(* Logix 5000 project; controller Seperator 1756-L85E rev 33.11; software revision 33.01; part 3 of 7 *)
(* tags used below, declared in another part *)
   Inp_RunFdbk : BOOL;   // Input Signal: RUN feedback from motor
   Inp_Sim : BOOL;   // 1=Simulate working motor; 0=Start/Stop/ Monitor actual motor
   Inp_OvrdCmd : DINT;   // Override Mode Command: 0=None, 1=Stop, 2=Start
   Cfg_HasRunFdbk : BOOL;   // 1=Motor provides run feedback
   Cfg_UseRunFdbk : BOOL;   // 1=Motor run feedback should be used for failure checking
   Cfg_AllowLocal : BOOL;   // 1=Allow Local Start/Stop without alarm, 0=Start/Stop from HMI/prog only
   Cfg_PCmdClear : ALIAS FOR Mode.Cfg_PCmdClear;
   Cfg_OperStopPrio : BOOL;   // 1=OCmd_Stop available in any mode, 0=OCmd_Stop only in Oper, Maint modes.
   Cfg_ShedOnFailToStart : BOOL;   // 1=Stop Motor and Alarm on Fail to Start; 0=Alarm only on Fail to Start
   PSet_Owner : DINT;   // Program Owner Request ID (non-zero) or Release (zero)
   PCmd_Start : BOOL;   // Program Command to Start Motor
   PCmd_Stop : BOOL;   // Program Command to Stop Motor
   PCmd_Reset : BOOL;   // Program Command to Reset all Alarms requiring Reset
   OCmd_Start : BOOL;   // Operator Command to Start Motor
   OCmd_Stop : BOOL;   // Operator Command to Stop Motor
   OCmd_Bypass : BOOL;   // Operator Command to Bypass all Bypassable Interlocks and Permissives
   OCmd_Check : BOOL;   // Operator Command to Check (not bypass) all Interlocks and Permissives
   MCmd_Disable : BOOL;   // Maintenance Command to Disable Motor
   MCmd_Enable : BOOL;   // Maintenance Command to Enable (allow to run) Motor
   OCmd_Reset : BOOL;   // Operator Command to Reset all Alarms requiring Reset
   OCmd_ResetAckAll : BOOL;   // Operator Command to Reset all Alarms and latched Shed conditions
   Out_Run : BOOL;   // 1=Run Motor, 0=Stop Motor
   Out_Start : BOOL;   // 1=Start Motor, 0=Motor left in current state
   Out_Stop : BOOL;   // 1=Stop Motor, 0=Motor left in current state
   Val_Cmd : SINT;   // Device Command 0=None, 1=Stop, 2=Start
   Val_Fdbk : SINT;   // Device Feedback 0=Stopped, 1=Running
   Val_Sts : SINT;   // Device Confirmed Sts 0=? 1=Stopped, 2=Running, 7=Stopping, 8=Starting, 33=Disabled
   Val_Fault : SINT;   // Device Fault Status 0=None, 16=Fail to Start, 17 = Fail to Stop, 32=I/O Fault, 34=Config Error
   Val_Owner : DINT;   // Current Object Owner ID (0=not owned)
   Val_Notify : SINT;   // Current Alarm Level and Acknowledgement (enumeration)
   Sts_Stopped : BOOL;   // 1=Motor requested to stop and is confirmed stopped
   Sts_Starting : BOOL;   // 1=Motor requested to run and awaiting run feedback
   Sts_Running : BOOL;   // 1=Motor requested to run and is confirmed running
   Sts_Stopping : BOOL;   // 1=Motor requested to stop and awaiting stopped feedback
   Sts_Available : BOOL;   // 1=Motor available for control by automation (Prog)
   Sts_Disabled : BOOL;   // 1=Motor is Disabled
   Sts_NotRdy : BOOL;   // 1=Motor is Not Ready to Run (independent of Mode)
   Sts_AlmInh : BOOL;   // 1=An Alarm is Shelved, Disabled or Suppressed: display icon
   Sts_Err : BOOL;   // 1=Error in Config: see detail bits for reason
   Sts_Hand : ALIAS FOR Mode.Sts_Hand;
   Sts_Maint : ALIAS FOR Mode.Sts_Maint;
   Sts_Ovrd : ALIAS FOR Mode.Sts_Ovrd;
   Sts_Prog : ALIAS FOR Mode.Sts_Prog;
   Sts_Oper : ALIAS FOR Mode.Sts_Oper;
   Sts_FailToStart : ALIAS FOR FailToStart.Inp;   // 1=Motor Failed to Start (one-shot)
   Sts_FailToStop : ALIAS FOR FailToStop.Inp;   // 1=Motor Failed to Stop
   Sts_IOFault : ALIAS FOR IOFault.Inp;   // I/O Comm Fault Status (0=OK, 1=Bad)
   Rdy_Start : BOOL;   // 1=Ready to receive OCmd_Start (enables HMI button)
   Rdy_Stop : BOOL;   // 1=Ready to receive OCmd_Stop (enables HMI button)
   Rdy_Reset : BOOL;   // 1=At least one Alarm or Latched Shed requires Reset
   Rdy_ResetAckAll : BOOL;   // 1=At least one Alarm or latched Shed condition requires Reset or Ack
   P_Motor : BOOL;   // Unique Parameter Name for auto - discovery
   Mode : P_Mode;   // Motor Mode Selection
   IOFault : P_Alarm;   // I/O Fault Alarm
   IntlkTrip : P_Alarm;   // Interlock Trip Alarm
   FailToStop : P_Alarm;   // Motor Failed to Stop Alarm
   FailToStart : P_Alarm;   // Motor Failed to Start Alarm
   Wrk_Run : BOOL;   // 1=Motor should be "running", 0=should be "stopped"
   Wrk_SimRunT : TIMER;   // Simulation Delay until Running
   Wrk_StopT : TIMER;   // Stop Check Timer
   Wrk_StartT : TIMER;   // Start Check Timer
   Wrk_SimStopT : TIMER;   // Simulation Delay until Stopped
   Wrk_RunFdbk : BOOL;   // Run Feedback based on mode, simulation, etc. 1=running
   Wrk_Notify : DINT;   // Buffer for building Val_Notify
   Wrk_Cmd : SINT;   // Buffer for building Val_Cmd
   Wrk_Sts : SINT;   // Buffer for building Val_Sts
   Wrk_Fault : SINT;   // Buffer for building Val_Fault
   Wrk_Retrigger : BOOL;   // Maint Start issued while running or Stop while stopped
   Wrk_FailToStart : BOOL;   // Fail to Start Fault (latched) stops motor and requires reset
   Wrk_IOFault : BOOL;   // I/O Fault (latched) stops motor and requires reset
   Starting : SFC_STEP;
   Stopped : SFC_STEP;
   Stopping : SFC_STEP;
(* P_Motor, continued *)

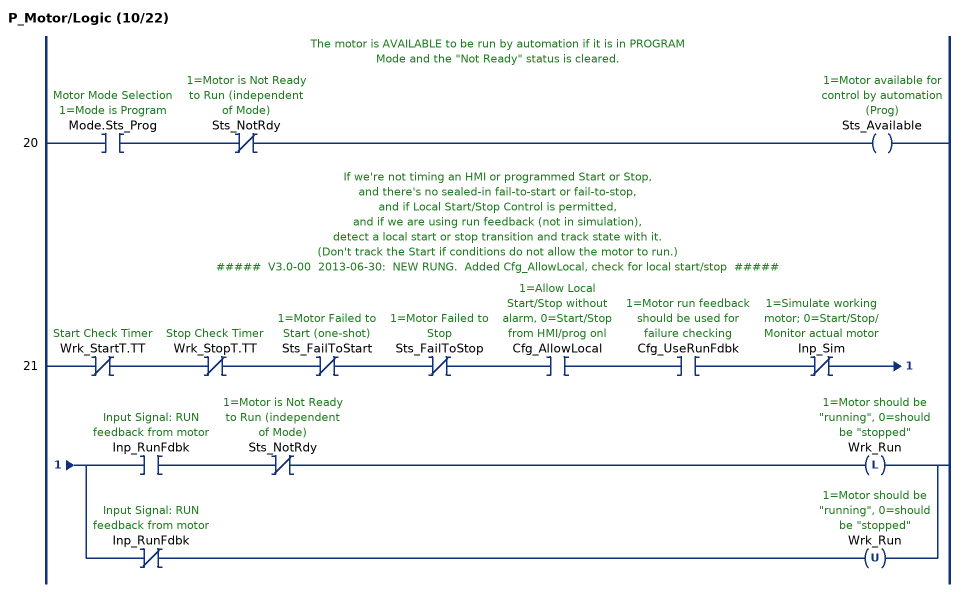
   // The motor is AVAILABLE to be run by automation if it is in PROGRAM
   // Mode and the "Not Ready" status is cleared.
   20: XIC(Mode.Sts_Prog)XIO(Sts_NotRdy)OTE(Sts_Available);
   // If we're not timing an HMI or programmed Start or Stop,
   // and there's no sealed-in fail-to-start or fail-to-stop,
   // and if Local Start/Stop Control is permitted,
   // and if we are using run feedback (not in simulation),
   // detect a local start or stop transition and track state with it.
   // (Don't track the Start if conditions do not allow the motor to run.)
   // #####  V3.0-00  2013-06-30:  NEW RUNG.  Added Cfg_AllowLocal, check for local start/stop  #####
   21: XIO(Wrk_StartT.TT)XIO(Wrk_StopT.TT)XIO(Sts_FailToStart)XIO(Sts_FailToStop)XIC(Cfg_AllowLocal)XIC(Cfg_UseRunFdbk)XIO(Inp_Sim)[XIC(Inp_RunFdbk) XIO(Sts_NotRdy) OTL(Wrk_Run) ,XIO(Inp_RunFdbk) OTU(Wrk_Run) ];
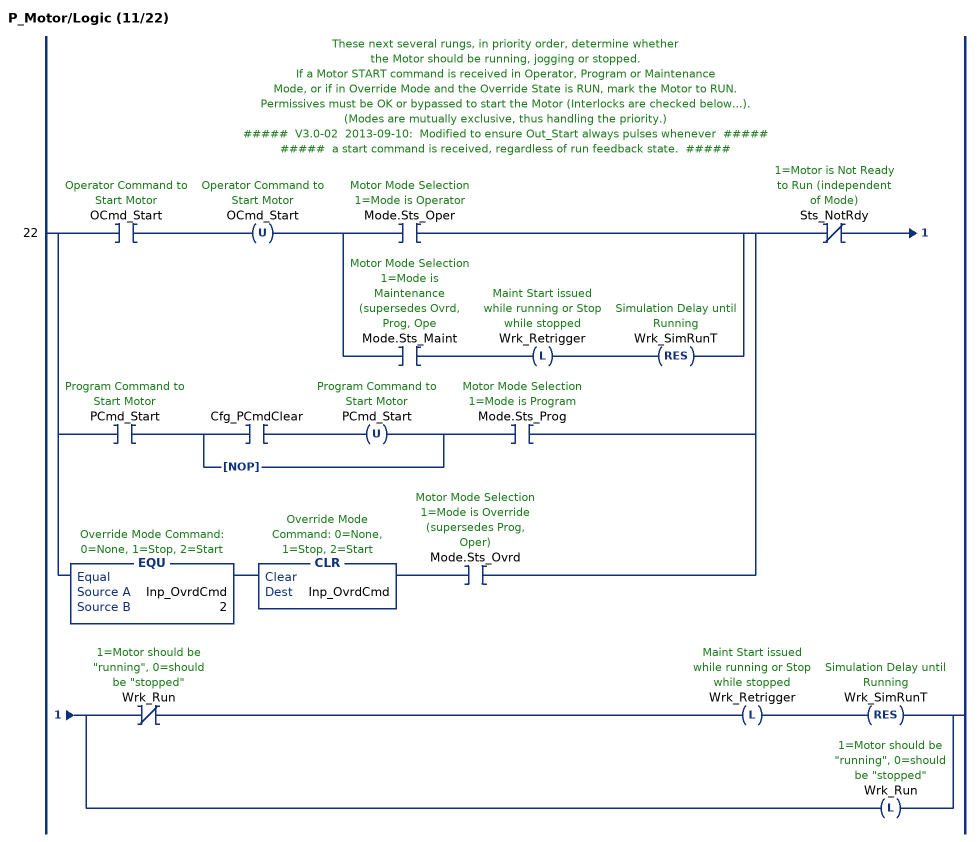
   // These next several rungs, in priority order, determine whether
   // the Motor should be running, jogging or stopped.
   // If a Motor START command is received in Operator, Program or Maintenance
   // Mode, or if in Override Mode and the Override State is RUN, mark the Motor to RUN.
   // Permissives must be OK or bypassed to start the Motor (Interlocks are checked below...).
   // (Modes are mutually exclusive, thus handling the priority.)
   // #####  V3.0-02  2013-09-10:  Modified to ensure Out_Start always pulses whenever  #####
   // #####  a start command is received, regardless of run feedback state.  #####
   22: [XIC(OCmd_Start) OTU(OCmd_Start) [XIC(Mode.Sts_Oper) ,XIC(Mode.Sts_Maint) OTL(Wrk_Retrigger) RES(Wrk_SimRunT) ] ,XIC(PCmd_Start) [XIC(Cfg_PCmdClear) OTU(PCmd_Start) ,NOP() ] XIC(Mode.Sts_Prog) ,EQU(Inp_OvrdCmd,2) CLR(Inp_OvrdCmd) XIC(Mode.Sts_Ovrd) ]XIO(Sts_NotRdy)[XIO(Wrk_Run) OTL(Wrk_Retrigger) RES(Wrk_SimRunT) ,OTL(Wrk_Run) ];
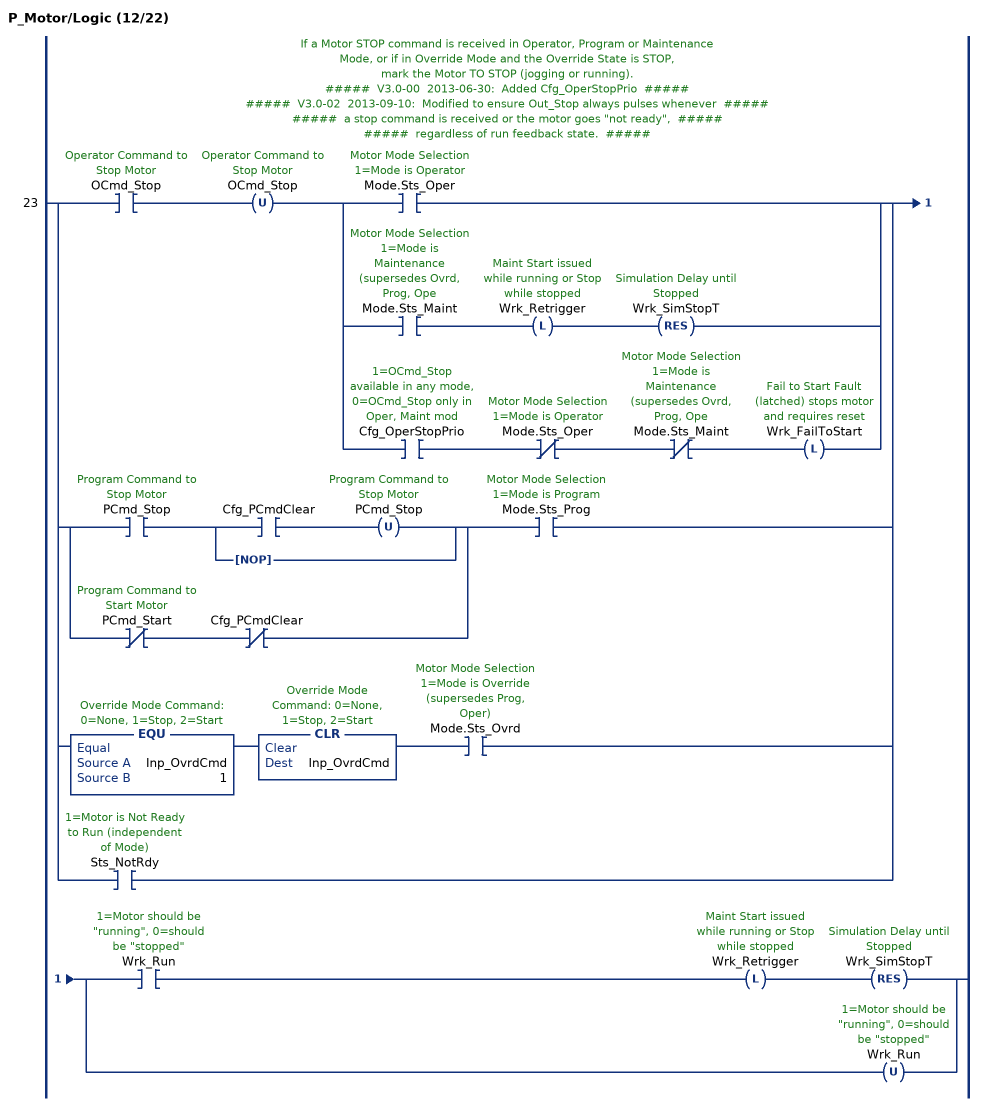
   // If a Motor STOP command is received in Operator, Program or Maintenance
   // Mode, or if in Override Mode and the Override State is STOP,
   // mark the Motor TO STOP (jogging or running).
   // #####  V3.0-00  2013-06-30:  Added Cfg_OperStopPrio  #####
   // #####  V3.0-02  2013-09-10:  Modified to ensure Out_Stop always pulses whenever  #####
   // #####  a stop command is received or the motor goes "not ready",  #####
   // #####  regardless of run feedback state.  #####
   23: [XIC(OCmd_Stop) OTU(OCmd_Stop) [XIC(Mode.Sts_Oper) ,XIC(Mode.Sts_Maint) OTL(Wrk_Retrigger) RES(Wrk_SimStopT) ,XIC(Cfg_OperStopPrio) XIO(Mode.Sts_Oper) XIO(Mode.Sts_Maint) OTL(Wrk_FailToStart) ] ,[XIC(PCmd_Stop) [XIC(Cfg_PCmdClear) OTU(PCmd_Stop) ,NOP() ] ,XIO(PCmd_Start) XIO(Cfg_PCmdClear) ] XIC(Mode.Sts_Prog) ,EQU(Inp_OvrdCmd,1) CLR(Inp_OvrdCmd) XIC(Mode.Sts_Ovrd) ,XIC(Sts_NotRdy) ][XIC(Wrk_Run) OTL(Wrk_Retrigger) RES(Wrk_SimStopT) ,OTU(Wrk_Run) ];
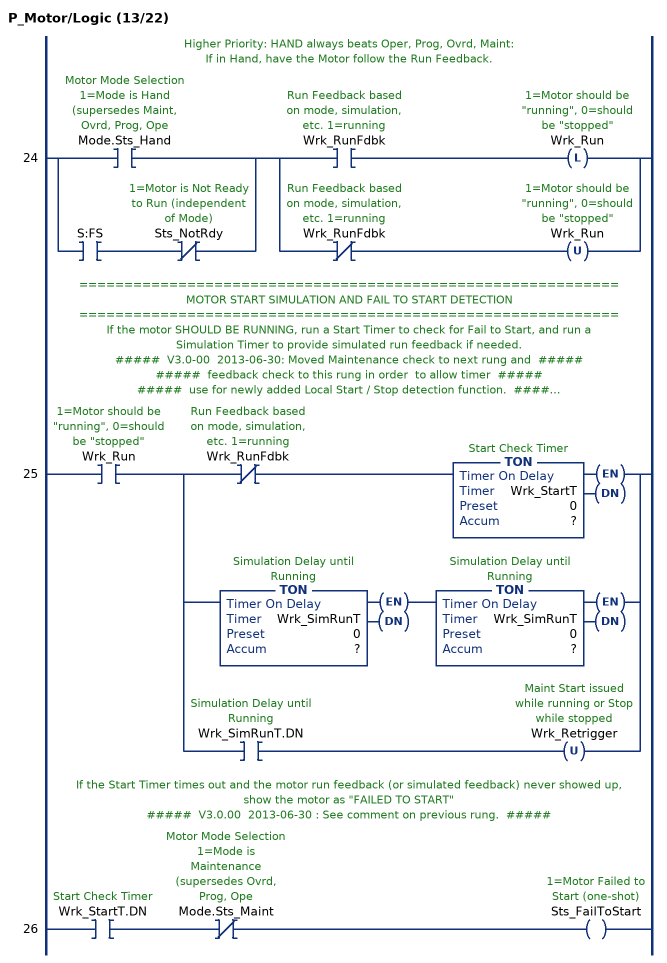
   // Higher Priority: HAND always beats Oper, Prog, Ovrd, Maint:
   // If in Hand, have the Motor follow the Run Feedback.
   24: [XIC(Mode.Sts_Hand) ,XIC(S:FS) XIO(Sts_NotRdy) ][XIC(Wrk_RunFdbk) OTL(Wrk_Run) ,XIO(Wrk_RunFdbk) OTU(Wrk_Run) ];
   // ============================================================
   // MOTOR START SIMULATION AND FAIL TO START DETECTION
   // ============================================================
   // If the motor SHOULD BE RUNNING, run a Start Timer to check for Fail to Start, and run a
   // Simulation Timer to provide simulated run feedback if needed.
   // #####  V3.0-00  2013-06-30: Moved Maintenance check to next rung and  #####
   // #####  feedback check to this rung in order  to allow timer  #####
   // #####  use for newly added Local Start / Stop detection function.  #####
   // @@@@@  The TON on the second branch is doubled to ensure it goes  @@@@@
   // @@@@@  the same scan it is enabled if its preset is zero.  @@@@@
   25: XIC(Wrk_Run)[XIO(Wrk_RunFdbk) TON(Wrk_StartT,?,?) ,TON(Wrk_SimRunT,?,?) TON(Wrk_SimRunT,?,?) ,XIC(Wrk_SimRunT.DN) OTU(Wrk_Retrigger) ];
   // If the Start Timer times out and the motor run feedback (or simulated feedback) never showed up,
   // show the motor as "FAILED TO START"
   // #####  V3.0.00  2013-06-30 : See comment on previous rung.  #####
   26: XIC(Wrk_StartT.DN)XIO(Mode.Sts_Maint)OTE(Sts_FailToStart);
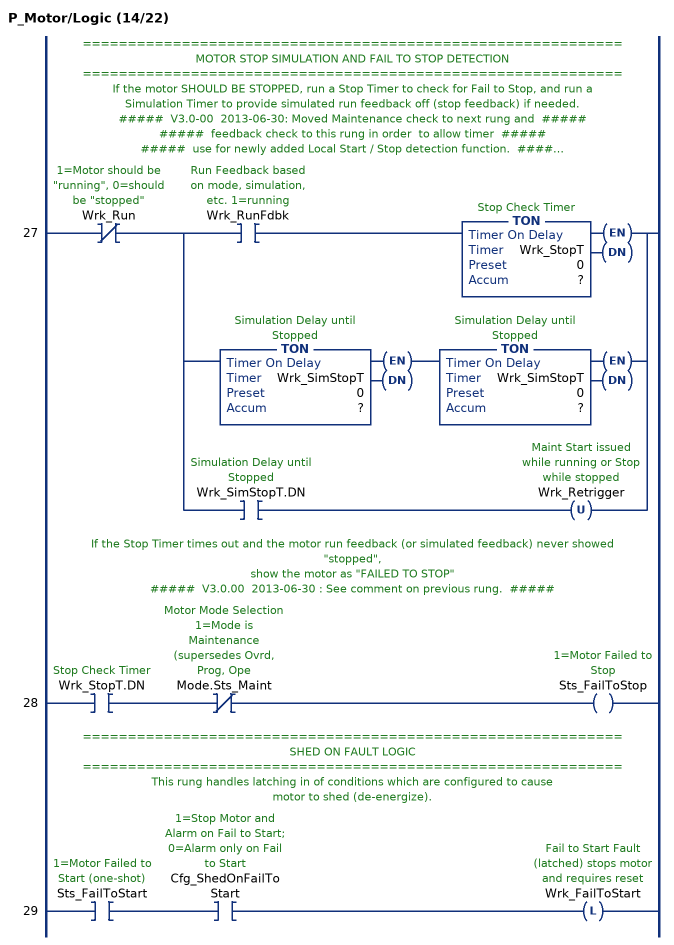
   // ============================================================
   // MOTOR STOP SIMULATION AND FAIL TO STOP DETECTION
   // ============================================================
   // If the motor SHOULD BE STOPPED, run a Stop Timer to check for Fail to Stop, and run a
   // Simulation Timer to provide simulated run feedback off (stop feedback) if needed.
   // #####  V3.0-00  2013-06-30: Moved Maintenance check to next rung and  #####
   // #####  feedback check to this rung in order  to allow timer  #####
   // #####  use for newly added Local Start / Stop detection function.  #####
   // @@@@@  The TON on the second branch is doubled to ensure it goes  @@@@@
   // @@@@@  the same scan it is enabled if its preset is zero.  @@@@@
   27: XIO(Wrk_Run)[XIC(Wrk_RunFdbk) TON(Wrk_StopT,?,?) ,TON(Wrk_SimStopT,?,?) TON(Wrk_SimStopT,?,?) ,XIC(Wrk_SimStopT.DN) OTU(Wrk_Retrigger) ];
   // If the Stop Timer times out and the motor run feedback (or simulated feedback) never showed "stopped",
   // show the motor as "FAILED TO STOP"
   // #####  V3.0.00  2013-06-30 : See comment on previous rung.  #####
   28: XIC(Wrk_StopT.DN)XIO(Mode.Sts_Maint)OTE(Sts_FailToStop);
   // ============================================================
   // SHED ON FAULT LOGIC
   // ============================================================
   // This rung handles latching in of conditions which are configured to cause
   // motor to shed (de-energize).
   29: XIC(Sts_FailToStart)XIC(Cfg_ShedOnFailToStart)OTL(Wrk_FailToStart);
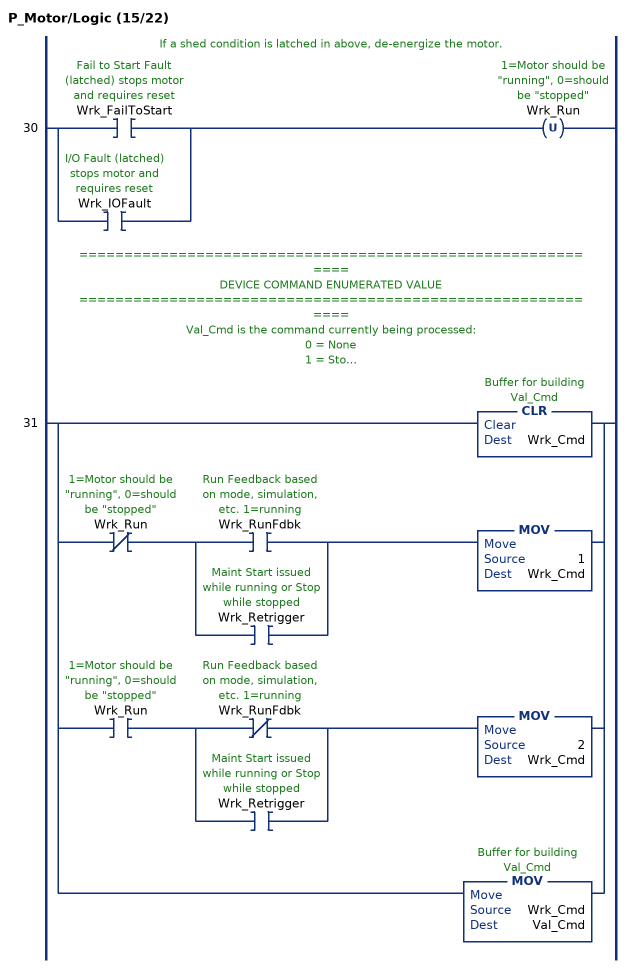
   // If a shed condition is latched in above, de-energize the motor.
   30: [XIC(Wrk_FailToStart) ,XIC(Wrk_IOFault) ]OTU(Wrk_Run);
   // ============================================================
   // DEVICE COMMAND ENUMERATED VALUE
   // ============================================================
   // Val_Cmd is the command currently being processed:
   // 0 = None
   // 1 = Stop
   // 2 = Start
   31: [CLR(Wrk_Cmd) ,XIO(Wrk_Run) [XIC(Wrk_RunFdbk) ,XIC(Wrk_Retrigger) ] MOV(1,Wrk_Cmd) ,XIC(Wrk_Run) [XIO(Wrk_RunFdbk) ,XIC(Wrk_Retrigger) ] MOV(2,Wrk_Cmd) ,MOV(Wrk_Cmd,Val_Cmd) ];
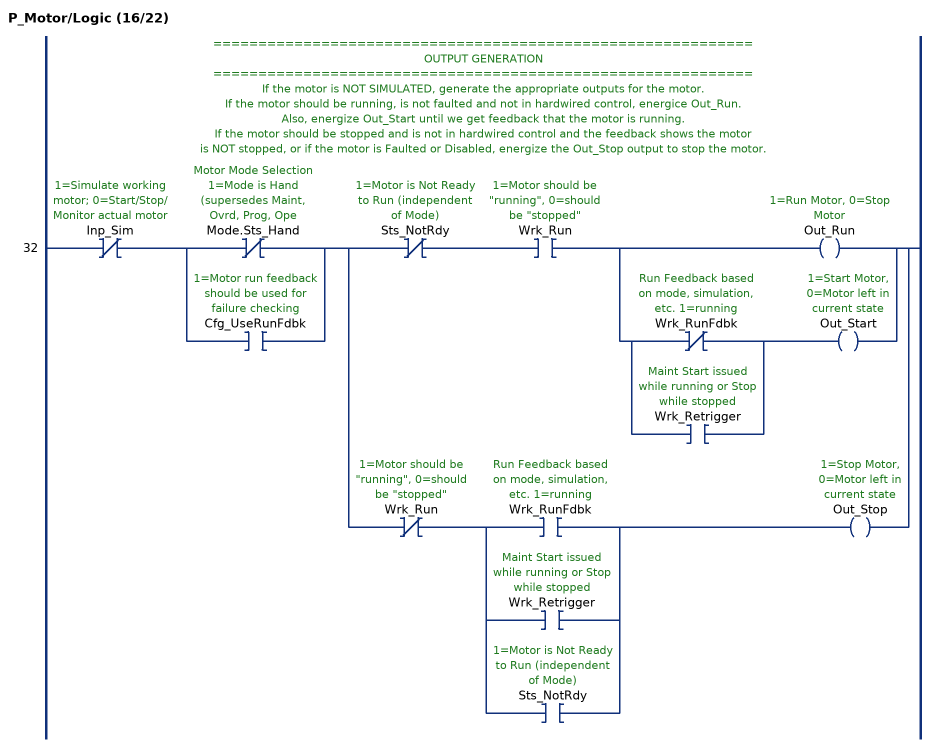
   // ============================================================
   // OUTPUT GENERATION
   // ============================================================
   // If the motor is NOT SIMULATED, generate the appropriate outputs for the motor.
   // If the motor should be running, is not faulted and not in hardwired control, energice Out_Run.
   // Also, energize Out_Start until we get feedback that the motor is running.
   // If the motor should be stopped and is not in hardwired control and the feedback shows the motor
   // is NOT stopped, or if the motor is Faulted or Disabled, energize the Out_Stop output to stop the motor.
   32: XIO(Inp_Sim)[XIO(Mode.Sts_Hand) ,XIC(Cfg_UseRunFdbk) ][XIO(Sts_NotRdy) XIC(Wrk_Run) [OTE(Out_Run) ,[XIO(Wrk_RunFdbk) ,XIC(Wrk_Retrigger) ] OTE(Out_Start) ] ,XIO(Wrk_Run) [XIC(Wrk_RunFdbk) ,XIC(Wrk_Retrigger) ,XIC(Sts_NotRdy) ] OTE(Out_Stop) ];
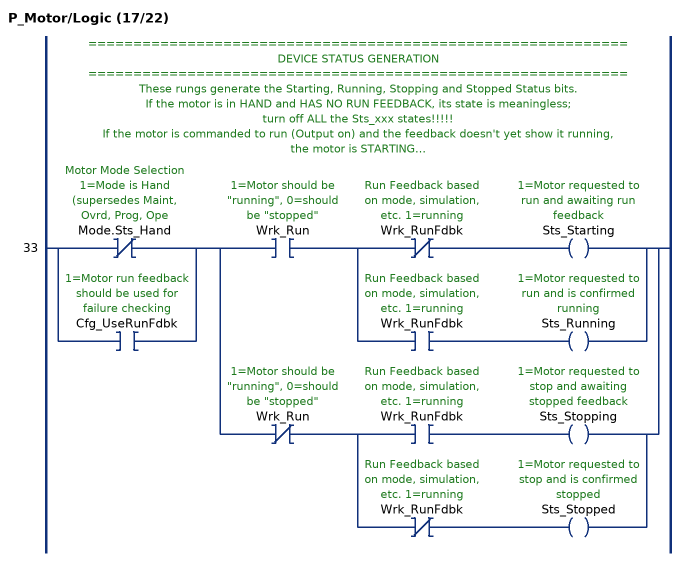
   // ============================================================
   // DEVICE STATUS GENERATION
   // ============================================================
   // These rungs generate the Starting, Running, Stopping and Stopped Status bits.
   // If the motor is in HAND and HAS NO RUN FEEDBACK, its state is meaningless;
   // turn off ALL the Sts_xxx states!!!!!
   // If the motor is commanded to run (Output on) and the feedback doesn't yet show it running,
   // the motor is STARTING.
   // If the motor is commanded to run (Output on) and the feedback shows it running,
   // the motor is RUNNING.
   // If the motor is commanded to stoop (Output off) and the feedback still shows it running,
   // the motor is STOPPING.
   // If the motor is commanded to stop (Output off) and the feedback shows it has stopped,
   // the motor is STOPPED.
   33: [XIO(Mode.Sts_Hand) ,XIC(Cfg_UseRunFdbk) ][XIC(Wrk_Run) [XIO(Wrk_RunFdbk) OTE(Sts_Starting) ,XIC(Wrk_RunFdbk) OTE(Sts_Running) ] ,XIO(Wrk_Run) [XIC(Wrk_RunFdbk) OTE(Sts_Stopping) ,XIO(Wrk_RunFdbk) OTE(Sts_Stopped) ] ];
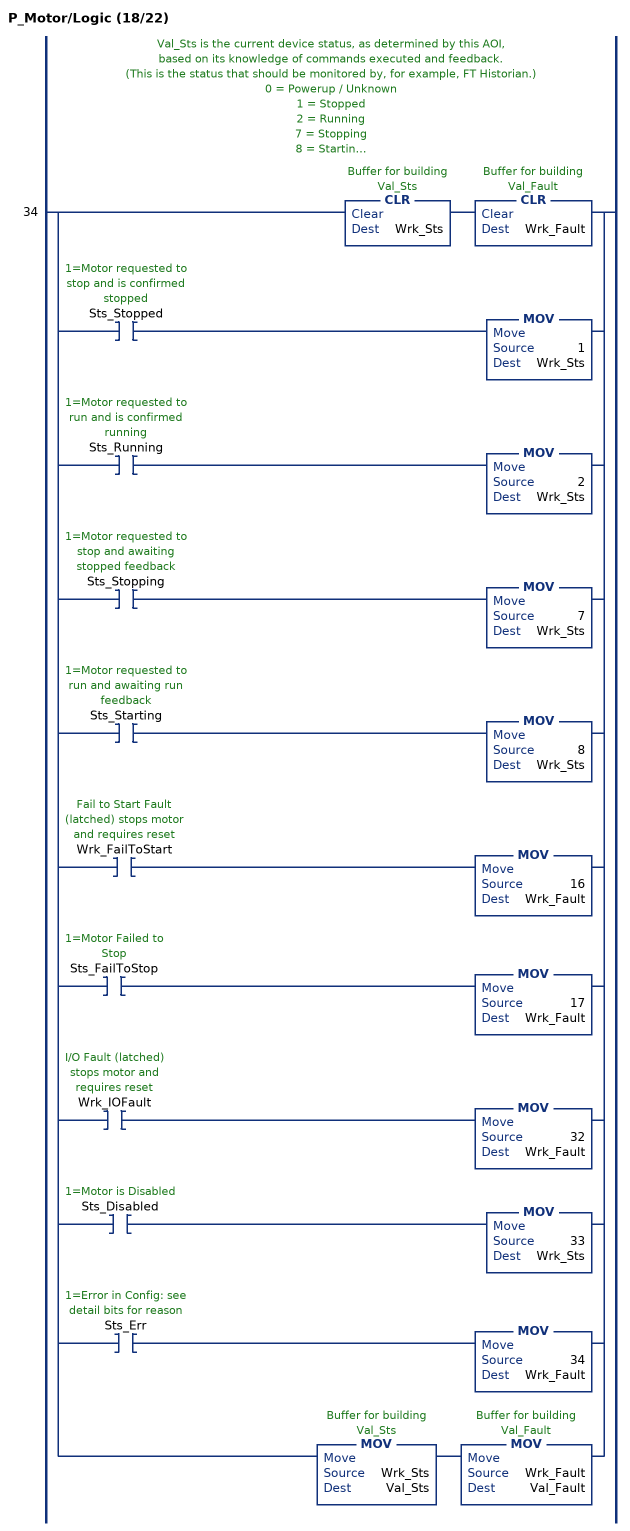
   // Val_Sts is the current device status, as determined by this AOI,
   // based on its knowledge of commands executed and feedback.
   // (This is the status that should be monitored by, for example, FT Historian.)
   // 0 = Powerup / Unknown
   // 1 = Stopped
   // 2 = Running
   // 7 = Stopping
   // 8 = Starting
   // 33 = Device Disabled
   // Val_Fault is the current device fault status, as determined by this AOI,
   // based on its knowledge of commands executed and feedback.
   // (This is the fault status that should be monitored by, for example, FT Historian.)
   // 0 = None
   // 16 = Fail to Start
   // 17 = Fail to Stop
   // 32 = I/O Fault (from Input)
   // 34 = Configuration Error
   34: [CLR(Wrk_Sts) CLR(Wrk_Fault) ,XIC(Sts_Stopped) MOV(1,Wrk_Sts) ,XIC(Sts_Running) MOV(2,Wrk_Sts) ,XIC(Sts_Stopping) MOV(7,Wrk_Sts) ,XIC(Sts_Starting) MOV(8,Wrk_Sts) ,XIC(Wrk_FailToStart) MOV(16,Wrk_Fault) ,XIC(Sts_FailToStop) MOV(17,Wrk_Fault) ,XIC(Wrk_IOFault) MOV(32,Wrk_Fault) ,XIC(Sts_Disabled) MOV(33,Wrk_Sts) ,XIC(Sts_Err) MOV(34,Wrk_Fault) ,MOV(Wrk_Sts,Val_Sts) MOV(Wrk_Fault,Val_Fault) ];
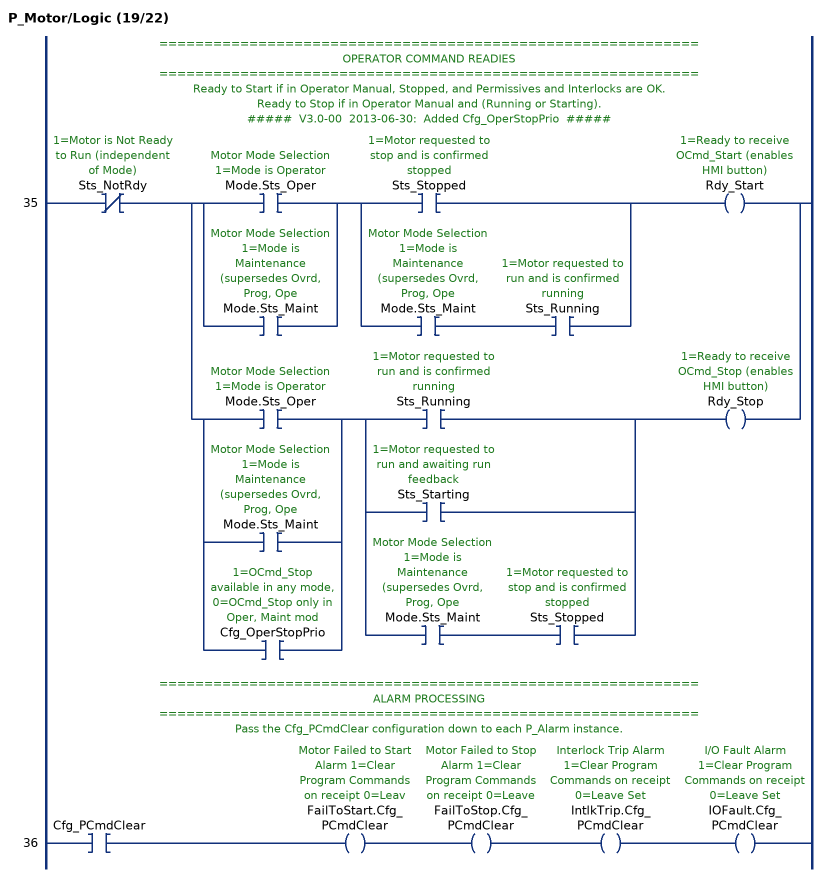
   // ============================================================
   // OPERATOR COMMAND READIES
   // ============================================================
   // Ready to Start if in Operator Manual, Stopped, and Permissives and Interlocks are OK.
   // Ready to Stop if in Operator Manual and (Running or Starting).
   // #####  V3.0-00  2013-06-30:  Added Cfg_OperStopPrio  #####
   35: XIO(Sts_NotRdy)[[XIC(Mode.Sts_Oper) ,XIC(Mode.Sts_Maint) ] [XIC(Sts_Stopped) ,XIC(Mode.Sts_Maint) XIC(Sts_Running) ] OTE(Rdy_Start) ,[XIC(Mode.Sts_Oper) ,XIC(Mode.Sts_Maint) ,XIC(Cfg_OperStopPrio) ] [XIC(Sts_Running) ,XIC(Sts_Starting) ,XIC(Mode.Sts_Maint) XIC(Sts_Stopped) ] OTE(Rdy_Stop) ];
   // ============================================================
   // ALARM PROCESSING
   // ============================================================
   // Pass the Cfg_PCmdClear configuration down to each P_Alarm instance.
   36: XIC(Cfg_PCmdClear)OTE(FailToStart.Cfg_PCmdClear)OTE(FailToStop.Cfg_PCmdClear)OTE(IntlkTrip.Cfg_PCmdClear)OTE(IOFault.Cfg_PCmdClear);
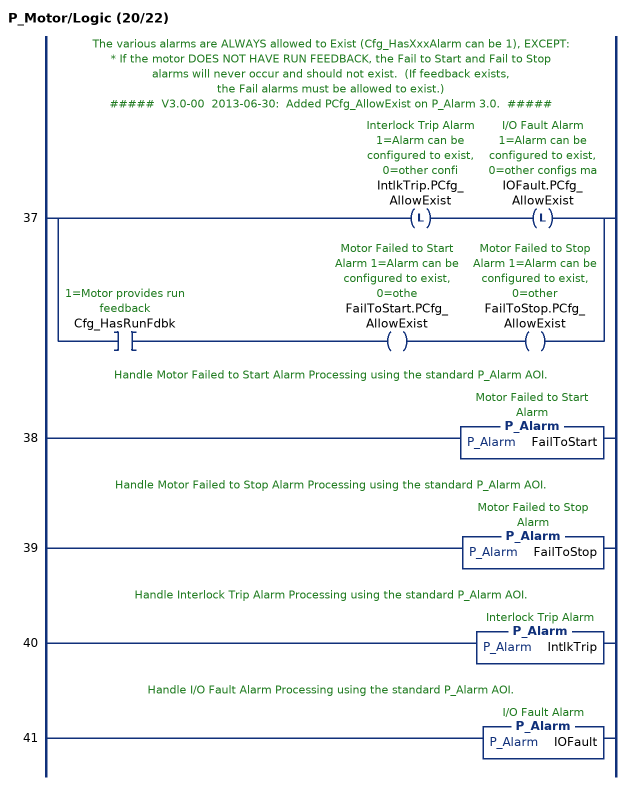
   // The various alarms are ALWAYS allowed to Exist (Cfg_HasXxxAlarm can be 1), EXCEPT:
   // * If the motor DOES NOT HAVE RUN FEEDBACK, the Fail to Start and Fail to Stop
   // alarms will never occur and should not exist.  (If feedback exists,
   // the Fail alarms must be allowed to exist.)
   // #####  V3.0-00  2013-06-30:  Added PCfg_AllowExist on P_Alarm 3.0.  #####
   37: [OTL(IntlkTrip.PCfg_AllowExist) OTL(IOFault.PCfg_AllowExist) ,XIC(Cfg_HasRunFdbk) OTE(FailToStart.PCfg_AllowExist) OTE(FailToStop.PCfg_AllowExist) ];
   // Handle Motor Failed to Start Alarm Processing using the standard P_Alarm AOI.
   38: P_Alarm(FailToStart);
   // Handle Motor Failed to Stop Alarm Processing using the standard P_Alarm AOI.
   39: P_Alarm(FailToStop);
   // Handle Interlock Trip Alarm Processing using the standard P_Alarm AOI.
   40: P_Alarm(IntlkTrip);
   // Handle I/O Fault Alarm Processing using the standard P_Alarm AOI.
   41: P_Alarm(IOFault);
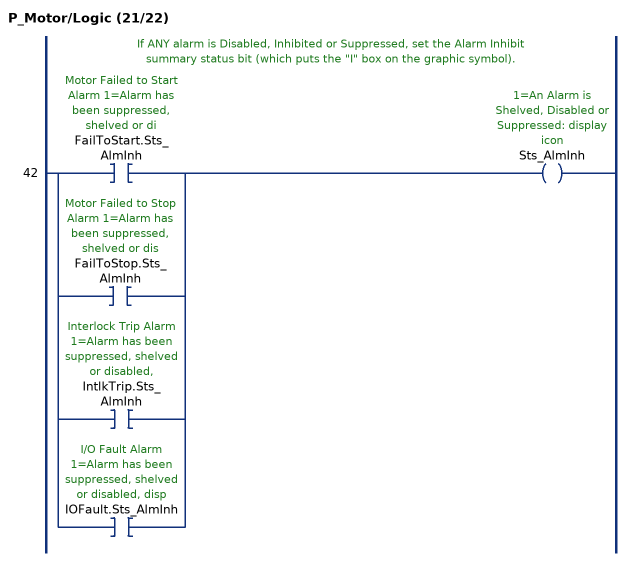
   // If ANY alarm is Disabled, Inhibited or Suppressed, set the Alarm Inhibit
   // summary status bit (which puts the "I" box on the graphic symbol).
   42: [XIC(FailToStart.Sts_AlmInh) ,XIC(FailToStop.Sts_AlmInh) ,XIC(IntlkTrip.Sts_AlmInh) ,XIC(IOFault.Sts_AlmInh) ]OTE(Sts_AlmInh);
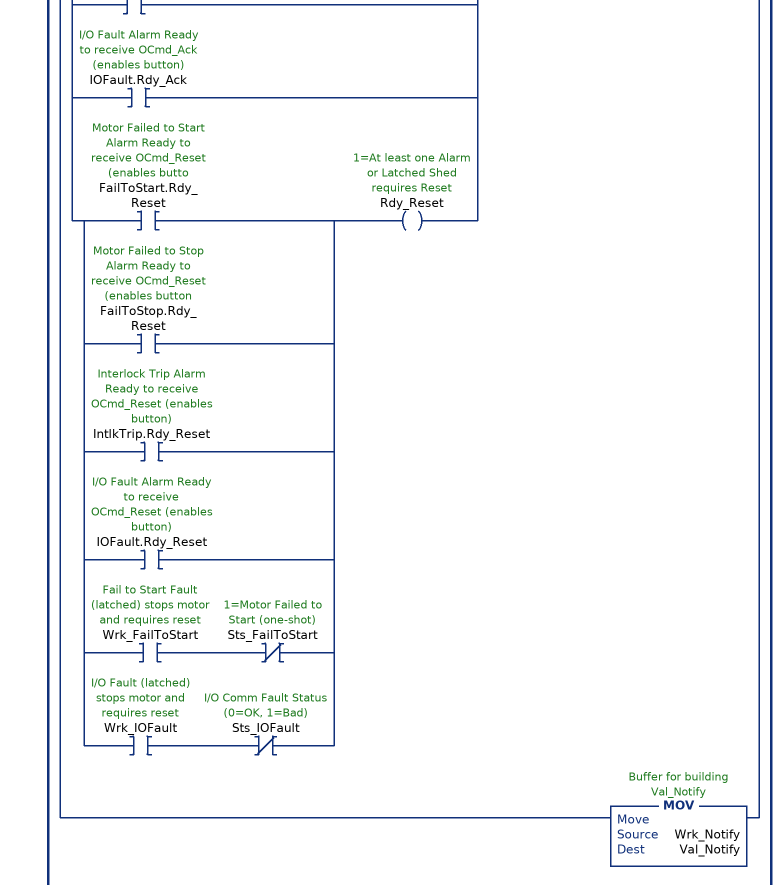
   // ============================================================
   // NOTIFICATION VALUE
   // ============================================================
   // Indicate the current alarm notification level as the max of any of the alarms,
   // and set the low-order bit for reset or ack required:
   // 0 = Not in alarm, acknowledged
   // 1 = Not in alarm, unacknowledged or reset required
   // 2 = Low severity alarm, acknowledged
   // 3 = Low severity alarm, unacknowledged
   // 4 = Medium severity alarm, acknowledged
   // 5 = Medium severity alarm, unacknowledged
   // 6 = High severity alarm, acknowledged
   // 7 = High severity alarm, unacknowledged
   // 8 = Highest severity alarm, acknowledged
   // 9 = Highest severity alarm, unacknowledged
   43: [CLR(Wrk_Notify) ,GRT(FailToStart.Val_Notify,Wrk_Notify) MOV(FailToStart.Val_Notify,Wrk_Notify) ,GRT(FailToStop.Val_Notify,Wrk_Notify) MOV(FailToStop.Val_Notify,Wrk_Notify) ,GRT(IntlkTrip.Val_Notify,Wrk_Notify) MOV(IntlkTrip.Val_Notify,Wrk_Notify) ,GRT(IOFault.Val_Notify,Wrk_Notify) MOV(IOFault.Val_Notify,Wrk_Notify) ,[[XIC(FailToStart.Rdy_Ack) ,XIC(FailToStop.Rdy_Ack) ,XIC(IntlkTrip.Rdy_Ack) ,XIC(IOFault.Rdy_Ack) ] ,[XIC(FailToStart.Rdy_Reset) ,XIC(FailToStop.Rdy_Reset) ,XIC(IntlkTrip.Rdy_Reset) ,XIC(IOFault.Rdy_Reset) ,XIC(Wrk_FailToStart) XIO(Sts_FailToStart) ,XIC(Wrk_IOFault) XIO(Sts_IOFault) ] OTE(Rdy_Reset) ] OTE(Rdy_ResetAckAll) OTE(Wrk_Notify.0) ,MOV(Wrk_Notify,Val_Notify) ];
END_ROUTINE

ROUTINE Prescan   (* ladder *)
// Clear Ownership, clear "lurking" Commands
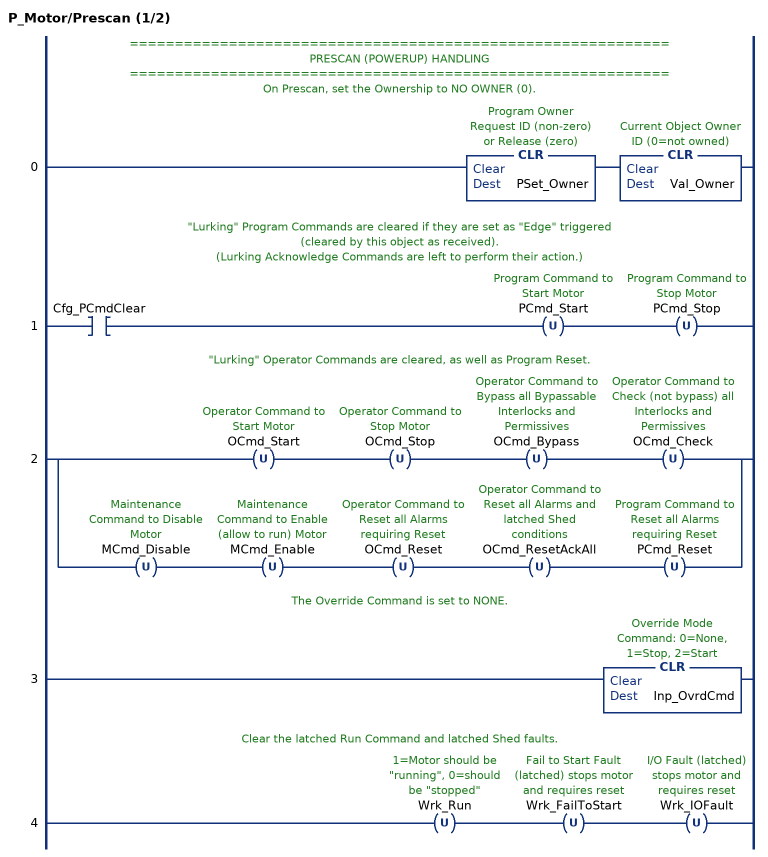
   // ============================================================
   // PRESCAN (POWERUP) HANDLING
   // ============================================================
   // On Prescan, set the Ownership to NO OWNER (0).
   0: CLR(PSet_Owner)CLR(Val_Owner);
   // "Lurking" Program Commands are cleared if they are set as "Edge" triggered
   // (cleared by this object as received).
   // (Lurking Acknowledge Commands are left to perform their action.)
   1: XIC(Cfg_PCmdClear)OTU(PCmd_Start)OTU(PCmd_Stop);
   // "Lurking" Operator Commands are cleared, as well as Program Reset.
   2: [OTU(OCmd_Start) OTU(OCmd_Stop) OTU(OCmd_Bypass) OTU(OCmd_Check) ,OTU(MCmd_Disable) OTU(MCmd_Enable) OTU(OCmd_Reset) OTU(OCmd_ResetAckAll) OTU(PCmd_Reset) ];
   // The Override Command is set to NONE.
   3: CLR(Inp_OvrdCmd);
   // Clear the latched Run Command and latched Shed faults.
   4: OTU(Wrk_Run)OTU(Wrk_FailToStart)OTU(Wrk_IOFault);
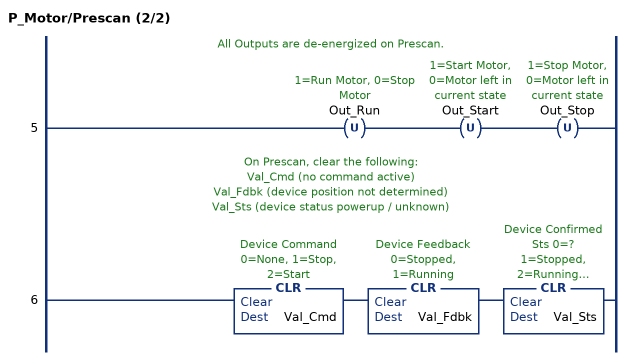
   // All Outputs are de-energized on Prescan.
   5: OTU(Out_Run)OTU(Out_Start)OTU(Out_Stop);
   // On Prescan, clear the following:
   // Val_Cmd (no command active)
   // Val_Fdbk (device position not determined)
   // Val_Sts (device status powerup / unknown)
   6: CLR(Val_Cmd)CLR(Val_Fdbk)CLR(Val_Sts);
END_ROUTINE
END_ADD_ON_INSTRUCTION

ADD_ON_INSTRUCTION RampUpDn   (* revision 1.0, vendor OGS, ExecutePrescan *)
VAR_INPUT
   CV : REAL; {required}
   Target : REAL; {required}
   Rate : REAL;
END_VAR
VAR_OUTPUT
   STS_RampDown : BOOL; {access Read Only, visible}
   STS_RampUp : BOOL; {access Read Only, visible}
   STS_Ramping : BOOL; {access Read Only, visible}
   STS_Dn : BOOL; {access Read Only, visible}
END_VAR
VAR_INPUT
   Time : REAL; {required}
END_VAR
VAR_OUTPUT
   output : REAL; {access Read Only, required}
END_VAR
VAR_INPUT
   CMD_Start : BOOL; {visible}
END_VAR
VAR
   Working : REAL;
   tmrSec : TIMER := (PRE := 1000);
   RatePerSec : REAL;
   ons : BOOL; {access None}
END_VAR

ROUTINE Logic   (* ladder *)
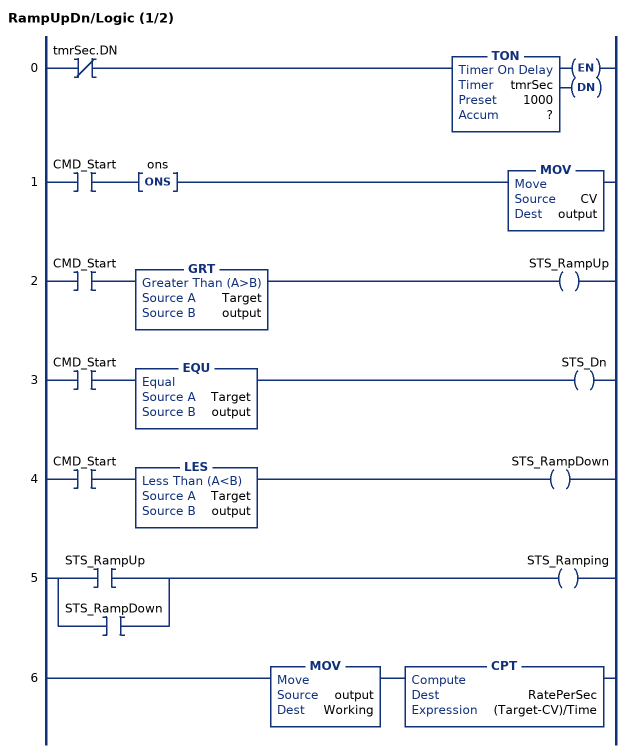
   0: XIO(tmrSec.DN)TON(tmrSec,?,?);
   1: XIC(CMD_Start)ONS(ons)MOV(CV,output);
   2: XIC(CMD_Start)GRT(Target,output)OTE(STS_RampUp);
   3: XIC(CMD_Start)EQU(Target,output)OTE(STS_Dn);
   4: XIC(CMD_Start)LES(Target,output)OTE(STS_RampDown);
   5: [XIC(STS_RampUp) ,XIC(STS_RampDown) ]OTE(STS_Ramping);
   6: MOV(output,Working)CPT(RatePerSec,(Target-CV)/Time);
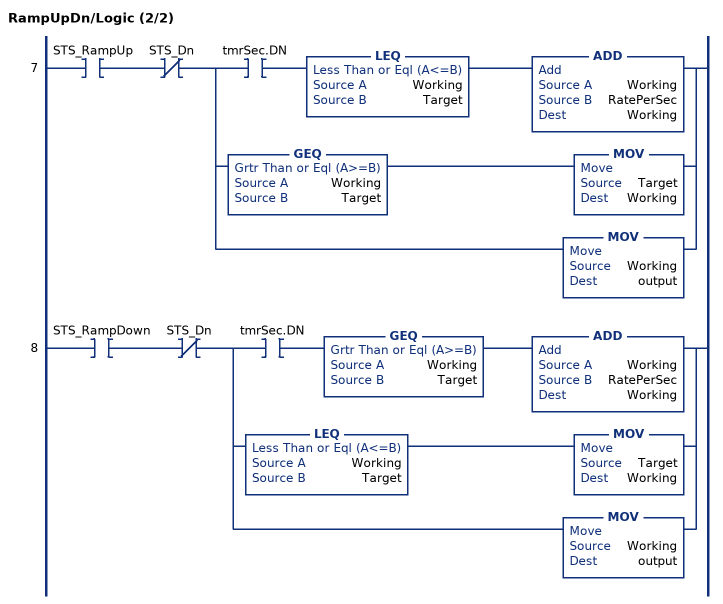
   7: XIC(STS_RampUp)XIO(STS_Dn)[XIC(tmrSec.DN) LEQ(Working,Target) ADD(Working,RatePerSec,Working) ,GEQ(Working,Target) MOV(Target,Working) ,MOV(Working,output) ];
   8: XIC(STS_RampDown)XIO(STS_Dn)[XIC(tmrSec.DN) GEQ(Working,Target) ADD(Working,RatePerSec,Working) ,LEQ(Working,Target) MOV(Target,Working) ,MOV(Working,output) ];
END_ROUTINE

ROUTINE Prescan   (* ladder *)
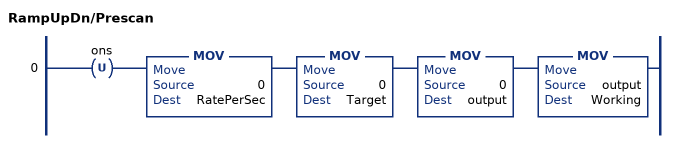
   0: OTU(ons)MOV(0,RatePerSec)MOV(0,Target)MOV(0,output)MOV(output,Working);
END_ROUTINE
END_ADD_ON_INSTRUCTION
